// TIA Portal project "Network_1.0" (V15.1)

(* hardware
DEVICE "S71500/ET200MP station_1"  S7-1500 station
   slot 0: "Rail_0"  Rack  6ES7 590-1***0-0AA0
   slot 1: "PLC_1"  CPU 1516-3 PN/DP  6ES7 516-3AN01-0AB0  V2.6
      slot 3: "CPU display_1"  6ES7591-1BA00-0AA0
   slot 2: "AI 8xU/I/RTD/TC ST_1"  AI 8xU/I/RTD/TC ST  6ES7 531-7KF00-0AB0  V2.2
   slot 3: "AQ 4xU/I ST_1"  AQ 4xU/I ST  6ES7 532-5HD00-0AB0  V2.2
   slot 4: "DI 32x24VDC HF_1"  DI 32x24VDC HF  6ES7 521-1BL00-0AB0  V2.1
   slot 5: "DQ 32x24VDC/0.5A HF_1"  DQ 32x24VDC/0.5A HF  6ES7 522-1BL01-0AB0  V1.1
DEVICE "S7-1200 station_1"  S7-1200 Station
   slot 0: "Rack_0"  S7-1200 Rack  Rack  V1.0
   slot 1: "PLC_2"  CPU 1215C DC/DC/DC  6ES7 215-1AG40-0XB0  V4.2
DEVICE "S7-1200 station_2"  S7-1200 Station
   slot 0: "Rack_0"  S7-1200 Rack  Rack  V1.0
   slot 1: "PLC_3"  CPU 1215C DC/DC/DC  6ES7 215-1AG40-0XB0  V4.2
DEVICE "HMI_1"  KTP400 Basic PN
   slot 0: "HMI_1"  KTP400 Basic PN  6AV2 123-2DB03-0AX0  15.1.0.0
   slot 1: "HMI_RT_1"  KTP400 Basic PN  6AV2 123-2DB03-0AX0  15.1.0.0
   slot 5: "HMI_1.IE_CP_1"  PROFINET Interface  15.0.1.0
      slot 1: "PROFINET Interface_1"  PROFINET Interface
         slot 1: "Port_1"  Port
DEVICE "HMI_2"  KTP400 Basic PN
   slot 0: "HMI_2"  KTP400 Basic PN  6AV2 123-2DB03-0AX0  15.1.0.0
   slot 1: "HMI_RT_2"  KTP400 Basic PN  6AV2 123-2DB03-0AX0  15.1.0.0
   slot 5: "HMI_2.IE_CP_1"  PROFINET Interface  15.0.1.0
      slot 1: "PROFINET Interface_1"  PROFINET Interface
         slot 1: "Port_1"  Port
DEVICE "HMI_3"  KTP400 Basic PN
   slot 0: "HMI_3"  KTP400 Basic PN  6AV2 123-2DB03-0AX0  15.1.0.0
   slot 1: "HMI_RT_3"  KTP400 Basic PN  6AV2 123-2DB03-0AX0  15.1.0.0
   slot 5: "HMI_3.IE_CP_1"  PROFINET Interface  15.0.1.0
      slot 1: "PROFINET Interface_1"  PROFINET Interface
         slot 1: "Port_1"  Port
DEVICE "SCALANCE X005"  SCALANCE X-Station
   slot 0: "SCALANCE X rack"  Rail
   slot 0: "Switch_1"  6GK5 005-0BA00-1AB2  V1.0
*)

// ===== PLC "PLC_1"  CPU 1516-3 PN/DP =====

VAR_GLOBAL   // PLC tag table "Default tag table"
   "H2_Bet" AT %Q9.6 : Bool;
   "S1_Bet" AT %I17.4 : Bool;
   "S2_Bet" AT %I17.5 : Bool;
   "S3_Bet" AT %I17.6 : Bool;
   "S4_Bet" AT %I17.7 : Bool;
   "PE_Bet" AT %I17.3 : Bool;
   "H1_Bet" AT %Q9.5 : Bool;
   "H3_Bet" AT %Q9.7 : Bool;
   "Clock_Byte" AT %MB20 : Byte;
   "Clock_10Hz" AT %M20.0 : Bool;
   "Clock_5Hz" AT %M20.1 : Bool;
   "Clock_2.5Hz" AT %M20.2 : Bool;
   "Clock_2Hz" AT %M20.3 : Bool;
   "Clock_1.25Hz" AT %M20.4 : Bool;
   "Clock_1Hz" AT %M20.5 : Bool;
   "Clock_0.625Hz" AT %M20.6 : Bool;
   "Clock_0.5Hz" AT %M20.7 : Bool;
END_VAR

VAR_GLOBAL   // PLC tag table "PLC_1"
   "Selector_HMI_1" AT %MW8 : UInt;
   "Selector_HMI_2" AT %MW10 : UInt;
   "Selector_HMI_3" AT %MW12 : UInt;
   "S1_HM1" AT %M3.0 : Bool;
   "S2_HM1" AT %M3.1 : Bool;
   "S3_HM1" AT %M3.2 : Bool;
   "S1_HM2" AT %M3.3 : Bool;
   "S2_HM2" AT %M3.4 : Bool;
   "S3_HM2" AT %M3.5 : Bool;
   "S1_HM3" AT %M3.6 : Bool;
   "S2_HM3" AT %M3.7 : Bool;
   "S3_HM3" AT %M4.0 : Bool;
   "S1_PL1" AT %M4.1 : Bool;
   "S2_PL1" AT %M4.2 : Bool;
   "S3_PL1" AT %M4.3 : Bool;
   "S1_PL2" AT %M4.4 : Bool;
   "S2_PL2" AT %M4.5 : Bool;
   "S3_PL2" AT %M4.6 : Bool;
   "S1_PL3" AT %M4.7 : Bool;
   "S2_PL3" AT %M5.0 : Bool;
   "S3_PL3" AT %M5.1 : Bool;
   "H1_PL1" AT %M5.2 : Bool;
   "H2_PL1" AT %M5.3 : Bool;
   "H3_PL1" AT %M5.4 : Bool;
   "H1_PL2" AT %M5.5 : Bool;
   "H2_PL2" AT %M5.6 : Bool;
   "H3_PL2" AT %M5.7 : Bool;
   "H1_PL3" AT %M6.0 : Bool;
   "H2_PL3" AT %M6.1 : Bool;
   "H3_PL3" AT %M6.2 : Bool;
   "H1_HM1" AT %M6.3 : Bool;
   "H2_HM1" AT %M6.4 : Bool;
   "H3_HM1" AT %M6.5 : Bool;
   "H1_HM2" AT %M6.6 : Bool;
   "H2_HM2" AT %M6.7 : Bool;
   "H3_HM2" AT %M7.0 : Bool;
   "H1_HM3" AT %M7.1 : Bool;
   "H2_HM3" AT %M7.2 : Bool;
   "H3_HM3" AT %M7.3 : Bool;
END_VAR

DATA_BLOCK "COMS_PLC"   // DB1
{ S7_Optimized_Access := 'FALSE' }
VERSION : 0.1
   VAR
      PLC2_H1 : Int;
      PLC2_H2 : Int;
      PLC2_H3 : Int;
      PLC3_H1 : Int;
      PLC3_H2 : Int;
      PLC3_H3 : Int;
      PLC1_S1 : Int;
      PLC1_S2 : Int;
      PLC1_S3 : Int;
      PLC2_S1 : Int;
      PLC2_S2 : Int;
      PLC2_S3 : Int;
      PLC3_S1 : Int;
      PLC3_S2 : Int;
      PLC3_S3 : Int;
   END_VAR
BEGIN
END_DATA_BLOCK

ORGANIZATION_BLOCK "Main"   // OB1, LAD, ProgramCycle
TITLE = "Main Program Sweep (Cycle)"
{ S7_Optimized_Access := 'TRUE' }
VERSION : 0.1
   VAR_INPUT
      Initial_Call : Bool;   // Initial call of this OB
      Remanence : Bool;   // =True, if remanent data are available
   END_VAR
BEGIN

REGION Network 1: Salidas a HMI1
   // Salidas a HMI Selector 1
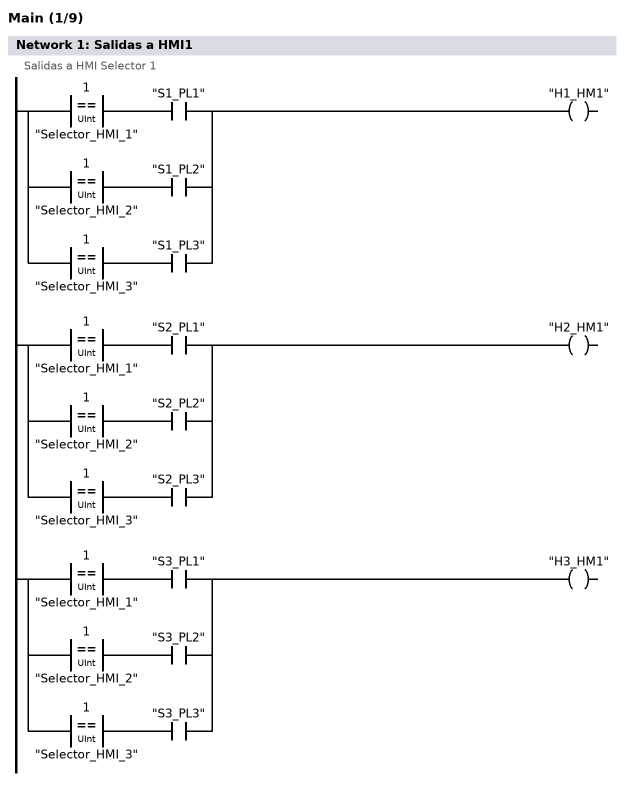
   RUNG wire#powerrail
      { S7_Templates := "SrcType := UInt" } EQ_Contact(in1 := 1, in2 := "Selector_HMI_1")
      Contact( "S1_PL1" )
      wire#w1
      Coil( "H1_HM1" )
   END_RUNG
   RUNG wire#powerrail
      { S7_Templates := "SrcType := UInt" } EQ_Contact(in1 := 1, in2 := "Selector_HMI_2")
      Contact( "S1_PL2" )
   END_RUNG wire#w1
   RUNG wire#powerrail
      { S7_Templates := "SrcType := UInt" } EQ_Contact(in1 := 1, in2 := "Selector_HMI_3")
      Contact( "S1_PL3" )
   END_RUNG wire#w1
   RUNG wire#powerrail
      { S7_Templates := "SrcType := UInt" } EQ_Contact(in1 := 1, in2 := "Selector_HMI_1")
      Contact( "S2_PL1" )
      wire#w2
      Coil( "H2_HM1" )
   END_RUNG
   RUNG wire#powerrail
      { S7_Templates := "SrcType := UInt" } EQ_Contact(in1 := 1, in2 := "Selector_HMI_2")
      Contact( "S2_PL2" )
   END_RUNG wire#w2
   RUNG wire#powerrail
      { S7_Templates := "SrcType := UInt" } EQ_Contact(in1 := 1, in2 := "Selector_HMI_3")
      Contact( "S2_PL3" )
   END_RUNG wire#w2
   RUNG wire#powerrail
      { S7_Templates := "SrcType := UInt" } EQ_Contact(in1 := 1, in2 := "Selector_HMI_1")
      Contact( "S3_PL1" )
      wire#w3
      Coil( "H3_HM1" )
   END_RUNG
   RUNG wire#powerrail
      { S7_Templates := "SrcType := UInt" } EQ_Contact(in1 := 1, in2 := "Selector_HMI_2")
      Contact( "S3_PL2" )
   END_RUNG wire#w3
   RUNG wire#powerrail
      { S7_Templates := "SrcType := UInt" } EQ_Contact(in1 := 1, in2 := "Selector_HMI_3")
      Contact( "S3_PL3" )
   END_RUNG wire#w3
   // the same network as SCL:
   "H1_HM1" := ((1 = "Selector_HMI_1") AND "S1_PL1") OR ((1 = "Selector_HMI_2") AND "S1_PL2") OR ((1 = "Selector_HMI_3") AND "S1_PL3");
   "H2_HM1" := ((1 = "Selector_HMI_1") AND "S2_PL1") OR ((1 = "Selector_HMI_2") AND "S2_PL2") OR ((1 = "Selector_HMI_3") AND "S2_PL3");
   "H3_HM1" := ((1 = "Selector_HMI_1") AND "S3_PL1") OR ((1 = "Selector_HMI_2") AND "S3_PL2") OR ((1 = "Selector_HMI_3") AND "S3_PL3");
END_REGION

REGION Network 2: Salidas a HMI2
   // Salidas a HMI Selector 1
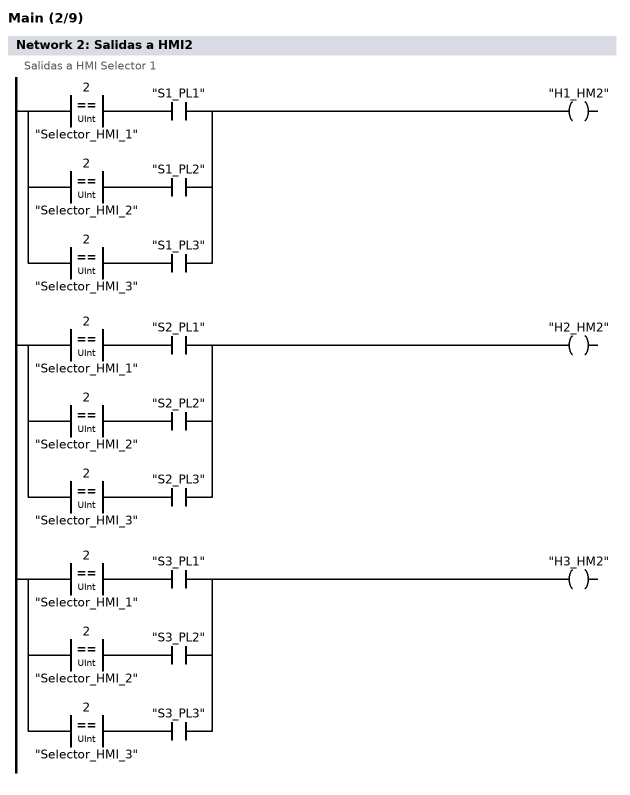
   RUNG wire#powerrail
      { S7_Templates := "SrcType := UInt" } EQ_Contact(in1 := 2, in2 := "Selector_HMI_1")
      Contact( "S1_PL1" )
      wire#w1
      Coil( "H1_HM2" )
   END_RUNG
   RUNG wire#powerrail
      { S7_Templates := "SrcType := UInt" } EQ_Contact(in1 := 2, in2 := "Selector_HMI_2")
      Contact( "S1_PL2" )
   END_RUNG wire#w1
   RUNG wire#powerrail
      { S7_Templates := "SrcType := UInt" } EQ_Contact(in1 := 2, in2 := "Selector_HMI_3")
      Contact( "S1_PL3" )
   END_RUNG wire#w1
   RUNG wire#powerrail
      { S7_Templates := "SrcType := UInt" } EQ_Contact(in1 := 2, in2 := "Selector_HMI_1")
      Contact( "S2_PL1" )
      wire#w2
      Coil( "H2_HM2" )
   END_RUNG
   RUNG wire#powerrail
      { S7_Templates := "SrcType := UInt" } EQ_Contact(in1 := 2, in2 := "Selector_HMI_2")
      Contact( "S2_PL2" )
   END_RUNG wire#w2
   RUNG wire#powerrail
      { S7_Templates := "SrcType := UInt" } EQ_Contact(in1 := 2, in2 := "Selector_HMI_3")
      Contact( "S2_PL3" )
   END_RUNG wire#w2
   RUNG wire#powerrail
      { S7_Templates := "SrcType := UInt" } EQ_Contact(in1 := 2, in2 := "Selector_HMI_1")
      Contact( "S3_PL1" )
      wire#w3
      Coil( "H3_HM2" )
   END_RUNG
   RUNG wire#powerrail
      { S7_Templates := "SrcType := UInt" } EQ_Contact(in1 := 2, in2 := "Selector_HMI_2")
      Contact( "S3_PL2" )
   END_RUNG wire#w3
   RUNG wire#powerrail
      { S7_Templates := "SrcType := UInt" } EQ_Contact(in1 := 2, in2 := "Selector_HMI_3")
      Contact( "S3_PL3" )
   END_RUNG wire#w3
   // the same network as SCL:
   "H1_HM2" := ((2 = "Selector_HMI_1") AND "S1_PL1") OR ((2 = "Selector_HMI_2") AND "S1_PL2") OR ((2 = "Selector_HMI_3") AND "S1_PL3");
   "H2_HM2" := ((2 = "Selector_HMI_1") AND "S2_PL1") OR ((2 = "Selector_HMI_2") AND "S2_PL2") OR ((2 = "Selector_HMI_3") AND "S2_PL3");
   "H3_HM2" := ((2 = "Selector_HMI_1") AND "S3_PL1") OR ((2 = "Selector_HMI_2") AND "S3_PL2") OR ((2 = "Selector_HMI_3") AND "S3_PL3");
END_REGION

REGION Network 3: Salidas a HMI3
   // Salidas a HMI Selector 1
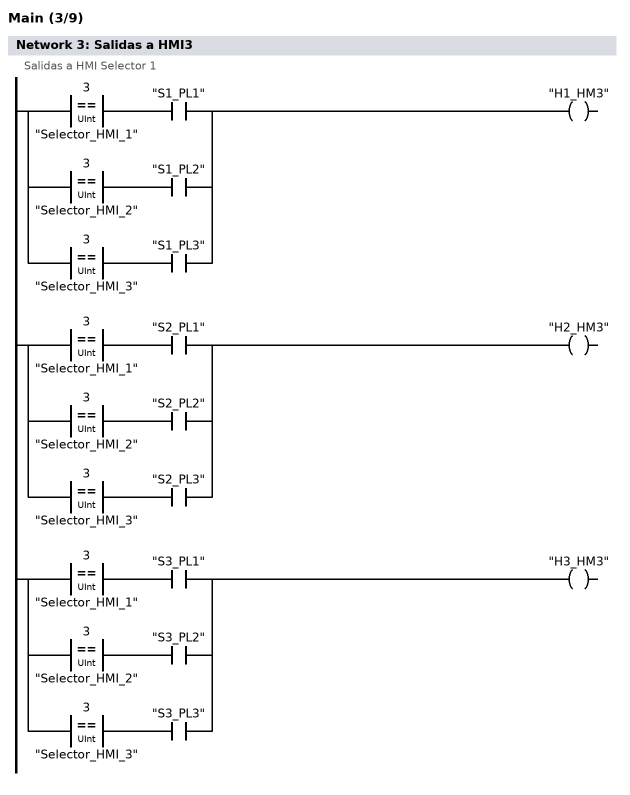
   RUNG wire#powerrail
      { S7_Templates := "SrcType := UInt" } EQ_Contact(in1 := 3, in2 := "Selector_HMI_1")
      Contact( "S1_PL1" )
      wire#w1
      Coil( "H1_HM3" )
   END_RUNG
   RUNG wire#powerrail
      { S7_Templates := "SrcType := UInt" } EQ_Contact(in1 := 3, in2 := "Selector_HMI_2")
      Contact( "S1_PL2" )
   END_RUNG wire#w1
   RUNG wire#powerrail
      { S7_Templates := "SrcType := UInt" } EQ_Contact(in1 := 3, in2 := "Selector_HMI_3")
      Contact( "S1_PL3" )
   END_RUNG wire#w1
   RUNG wire#powerrail
      { S7_Templates := "SrcType := UInt" } EQ_Contact(in1 := 3, in2 := "Selector_HMI_1")
      Contact( "S2_PL1" )
      wire#w2
      Coil( "H2_HM3" )
   END_RUNG
   RUNG wire#powerrail
      { S7_Templates := "SrcType := UInt" } EQ_Contact(in1 := 3, in2 := "Selector_HMI_2")
      Contact( "S2_PL2" )
   END_RUNG wire#w2
   RUNG wire#powerrail
      { S7_Templates := "SrcType := UInt" } EQ_Contact(in1 := 3, in2 := "Selector_HMI_3")
      Contact( "S2_PL3" )
   END_RUNG wire#w2
   RUNG wire#powerrail
      { S7_Templates := "SrcType := UInt" } EQ_Contact(in1 := 3, in2 := "Selector_HMI_1")
      Contact( "S3_PL1" )
      wire#w3
      Coil( "H3_HM3" )
   END_RUNG
   RUNG wire#powerrail
      { S7_Templates := "SrcType := UInt" } EQ_Contact(in1 := 3, in2 := "Selector_HMI_2")
      Contact( "S3_PL2" )
   END_RUNG wire#w3
   RUNG wire#powerrail
      { S7_Templates := "SrcType := UInt" } EQ_Contact(in1 := 3, in2 := "Selector_HMI_3")
      Contact( "S3_PL3" )
   END_RUNG wire#w3
   // the same network as SCL:
   "H1_HM3" := ((3 = "Selector_HMI_1") AND "S1_PL1") OR ((3 = "Selector_HMI_2") AND "S1_PL2") OR ((3 = "Selector_HMI_3") AND "S1_PL3");
   "H2_HM3" := ((3 = "Selector_HMI_1") AND "S2_PL1") OR ((3 = "Selector_HMI_2") AND "S2_PL2") OR ((3 = "Selector_HMI_3") AND "S2_PL3");
   "H3_HM3" := ((3 = "Selector_HMI_1") AND "S3_PL1") OR ((3 = "Selector_HMI_2") AND "S3_PL2") OR ((3 = "Selector_HMI_3") AND "S3_PL3");
END_REGION

REGION Network 4: Salidas a PLC1
   // Salidas a HMI Selector 1
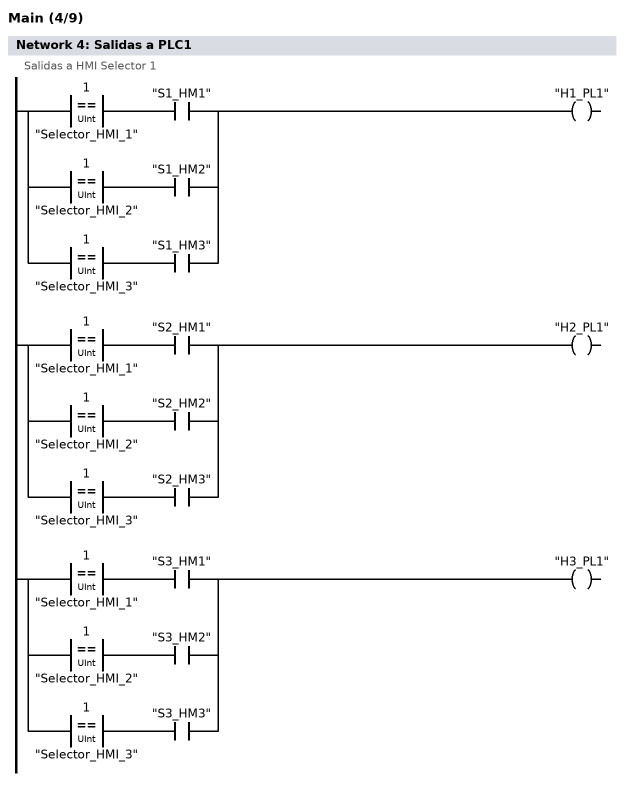
   RUNG wire#powerrail
      { S7_Templates := "SrcType := UInt" } EQ_Contact(in1 := 1, in2 := "Selector_HMI_1")
      Contact( "S1_HM1" )
      wire#w1
      Coil( "H1_PL1" )
   END_RUNG
   RUNG wire#powerrail
      { S7_Templates := "SrcType := UInt" } EQ_Contact(in1 := 1, in2 := "Selector_HMI_2")
      Contact( "S1_HM2" )
   END_RUNG wire#w1
   RUNG wire#powerrail
      { S7_Templates := "SrcType := UInt" } EQ_Contact(in1 := 1, in2 := "Selector_HMI_3")
      Contact( "S1_HM3" )
   END_RUNG wire#w1
   RUNG wire#powerrail
      { S7_Templates := "SrcType := UInt" } EQ_Contact(in1 := 1, in2 := "Selector_HMI_1")
      Contact( "S2_HM1" )
      wire#w2
      Coil( "H2_PL1" )
   END_RUNG
   RUNG wire#powerrail
      { S7_Templates := "SrcType := UInt" } EQ_Contact(in1 := 1, in2 := "Selector_HMI_2")
      Contact( "S2_HM2" )
   END_RUNG wire#w2
   RUNG wire#powerrail
      { S7_Templates := "SrcType := UInt" } EQ_Contact(in1 := 1, in2 := "Selector_HMI_3")
      Contact( "S2_HM3" )
   END_RUNG wire#w2
   RUNG wire#powerrail
      { S7_Templates := "SrcType := UInt" } EQ_Contact(in1 := 1, in2 := "Selector_HMI_1")
      Contact( "S3_HM1" )
      wire#w3
      Coil( "H3_PL1" )
   END_RUNG
   RUNG wire#powerrail
      { S7_Templates := "SrcType := UInt" } EQ_Contact(in1 := 1, in2 := "Selector_HMI_2")
      Contact( "S3_HM2" )
   END_RUNG wire#w3
   RUNG wire#powerrail
      { S7_Templates := "SrcType := UInt" } EQ_Contact(in1 := 1, in2 := "Selector_HMI_3")
      Contact( "S3_HM3" )
   END_RUNG wire#w3
   // the same network as SCL:
   "H1_PL1" := ((1 = "Selector_HMI_1") AND "S1_HM1") OR ((1 = "Selector_HMI_2") AND "S1_HM2") OR ((1 = "Selector_HMI_3") AND "S1_HM3");
   "H2_PL1" := ((1 = "Selector_HMI_1") AND "S2_HM1") OR ((1 = "Selector_HMI_2") AND "S2_HM2") OR ((1 = "Selector_HMI_3") AND "S2_HM3");
   "H3_PL1" := ((1 = "Selector_HMI_1") AND "S3_HM1") OR ((1 = "Selector_HMI_2") AND "S3_HM2") OR ((1 = "Selector_HMI_3") AND "S3_HM3");
END_REGION

REGION Network 5: Salidas a PLC2
   // Salidas a HMI Selector 1
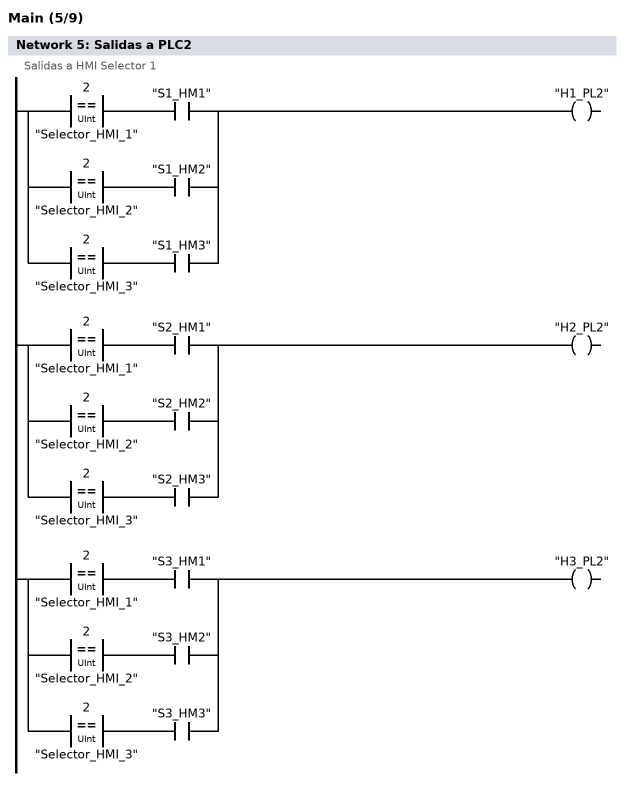
   RUNG wire#powerrail
      { S7_Templates := "SrcType := UInt" } EQ_Contact(in1 := 2, in2 := "Selector_HMI_1")
      Contact( "S1_HM1" )
      wire#w1
      Coil( "H1_PL2" )
   END_RUNG
   RUNG wire#powerrail
      { S7_Templates := "SrcType := UInt" } EQ_Contact(in1 := 2, in2 := "Selector_HMI_2")
      Contact( "S1_HM2" )
   END_RUNG wire#w1
   RUNG wire#powerrail
      { S7_Templates := "SrcType := UInt" } EQ_Contact(in1 := 2, in2 := "Selector_HMI_3")
      Contact( "S1_HM3" )
   END_RUNG wire#w1
   RUNG wire#powerrail
      { S7_Templates := "SrcType := UInt" } EQ_Contact(in1 := 2, in2 := "Selector_HMI_1")
      Contact( "S2_HM1" )
      wire#w2
      Coil( "H2_PL2" )
   END_RUNG
   RUNG wire#powerrail
      { S7_Templates := "SrcType := UInt" } EQ_Contact(in1 := 2, in2 := "Selector_HMI_2")
      Contact( "S2_HM2" )
   END_RUNG wire#w2
   RUNG wire#powerrail
      { S7_Templates := "SrcType := UInt" } EQ_Contact(in1 := 2, in2 := "Selector_HMI_3")
      Contact( "S2_HM3" )
   END_RUNG wire#w2
   RUNG wire#powerrail
      { S7_Templates := "SrcType := UInt" } EQ_Contact(in1 := 2, in2 := "Selector_HMI_1")
      Contact( "S3_HM1" )
      wire#w3
      Coil( "H3_PL2" )
   END_RUNG
   RUNG wire#powerrail
      { S7_Templates := "SrcType := UInt" } EQ_Contact(in1 := 2, in2 := "Selector_HMI_2")
      Contact( "S3_HM2" )
   END_RUNG wire#w3
   RUNG wire#powerrail
      { S7_Templates := "SrcType := UInt" } EQ_Contact(in1 := 2, in2 := "Selector_HMI_3")
      Contact( "S3_HM3" )
   END_RUNG wire#w3
   // the same network as SCL:
   "H1_PL2" := ((2 = "Selector_HMI_1") AND "S1_HM1") OR ((2 = "Selector_HMI_2") AND "S1_HM2") OR ((2 = "Selector_HMI_3") AND "S1_HM3");
   "H2_PL2" := ((2 = "Selector_HMI_1") AND "S2_HM1") OR ((2 = "Selector_HMI_2") AND "S2_HM2") OR ((2 = "Selector_HMI_3") AND "S2_HM3");
   "H3_PL2" := ((2 = "Selector_HMI_1") AND "S3_HM1") OR ((2 = "Selector_HMI_2") AND "S3_HM2") OR ((2 = "Selector_HMI_3") AND "S3_HM3");
END_REGION

REGION Network 6: Salidas a PLC3
   // Salidas a HMI Selector 1
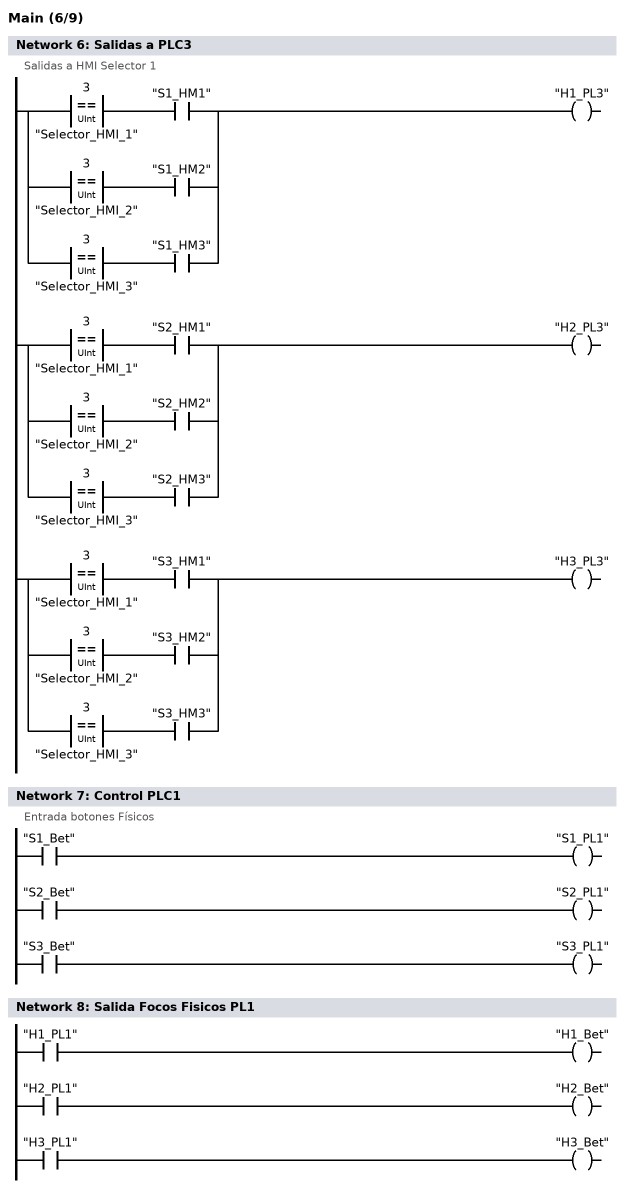
   RUNG wire#powerrail
      { S7_Templates := "SrcType := UInt" } EQ_Contact(in1 := 3, in2 := "Selector_HMI_1")
      Contact( "S1_HM1" )
      wire#w1
      Coil( "H1_PL3" )
   END_RUNG
   RUNG wire#powerrail
      { S7_Templates := "SrcType := UInt" } EQ_Contact(in1 := 3, in2 := "Selector_HMI_2")
      Contact( "S1_HM2" )
   END_RUNG wire#w1
   RUNG wire#powerrail
      { S7_Templates := "SrcType := UInt" } EQ_Contact(in1 := 3, in2 := "Selector_HMI_3")
      Contact( "S1_HM3" )
   END_RUNG wire#w1
   RUNG wire#powerrail
      { S7_Templates := "SrcType := UInt" } EQ_Contact(in1 := 3, in2 := "Selector_HMI_1")
      Contact( "S2_HM1" )
      wire#w2
      Coil( "H2_PL3" )
   END_RUNG
   RUNG wire#powerrail
      { S7_Templates := "SrcType := UInt" } EQ_Contact(in1 := 3, in2 := "Selector_HMI_2")
      Contact( "S2_HM2" )
   END_RUNG wire#w2
   RUNG wire#powerrail
      { S7_Templates := "SrcType := UInt" } EQ_Contact(in1 := 3, in2 := "Selector_HMI_3")
      Contact( "S2_HM3" )
   END_RUNG wire#w2
   RUNG wire#powerrail
      { S7_Templates := "SrcType := UInt" } EQ_Contact(in1 := 3, in2 := "Selector_HMI_1")
      Contact( "S3_HM1" )
      wire#w3
      Coil( "H3_PL3" )
   END_RUNG
   RUNG wire#powerrail
      { S7_Templates := "SrcType := UInt" } EQ_Contact(in1 := 3, in2 := "Selector_HMI_2")
      Contact( "S3_HM2" )
   END_RUNG wire#w3
   RUNG wire#powerrail
      { S7_Templates := "SrcType := UInt" } EQ_Contact(in1 := 3, in2 := "Selector_HMI_3")
      Contact( "S3_HM3" )
   END_RUNG wire#w3
   // the same network as SCL:
   "H1_PL3" := ((3 = "Selector_HMI_1") AND "S1_HM1") OR ((3 = "Selector_HMI_2") AND "S1_HM2") OR ((3 = "Selector_HMI_3") AND "S1_HM3");
   "H2_PL3" := ((3 = "Selector_HMI_1") AND "S2_HM1") OR ((3 = "Selector_HMI_2") AND "S2_HM2") OR ((3 = "Selector_HMI_3") AND "S2_HM3");
   "H3_PL3" := ((3 = "Selector_HMI_1") AND "S3_HM1") OR ((3 = "Selector_HMI_2") AND "S3_HM2") OR ((3 = "Selector_HMI_3") AND "S3_HM3");
END_REGION

REGION Network 7: Control PLC1
   // Entrada botones Físicos
   RUNG wire#powerrail
      Contact( "S1_Bet" )
      Coil( "S1_PL1" )
   END_RUNG
   RUNG wire#powerrail
      Contact( "S2_Bet" )
      Coil( "S2_PL1" )
   END_RUNG
   RUNG wire#powerrail
      Contact( "S3_Bet" )
      Coil( "S3_PL1" )
   END_RUNG
   // the same network as SCL:
   "S1_PL1" := "S1_Bet";
   "S2_PL1" := "S2_Bet";
   "S3_PL1" := "S3_Bet";
END_REGION

REGION Network 8: Salida Focos Fisicos PL1
   RUNG wire#powerrail
      Contact( "H1_PL1" )
      Coil( "H1_Bet" )
   END_RUNG
   RUNG wire#powerrail
      Contact( "H2_PL1" )
      Coil( "H2_Bet" )
   END_RUNG
   RUNG wire#powerrail
      Contact( "H3_PL1" )
      Coil( "H3_Bet" )
   END_RUNG
   // the same network as SCL:
   "H1_Bet" := "H1_PL1";
   "H2_Bet" := "H2_PL1";
   "H3_Bet" := "H3_PL1";
END_REGION

REGION Network 9: LECTURAS PLC
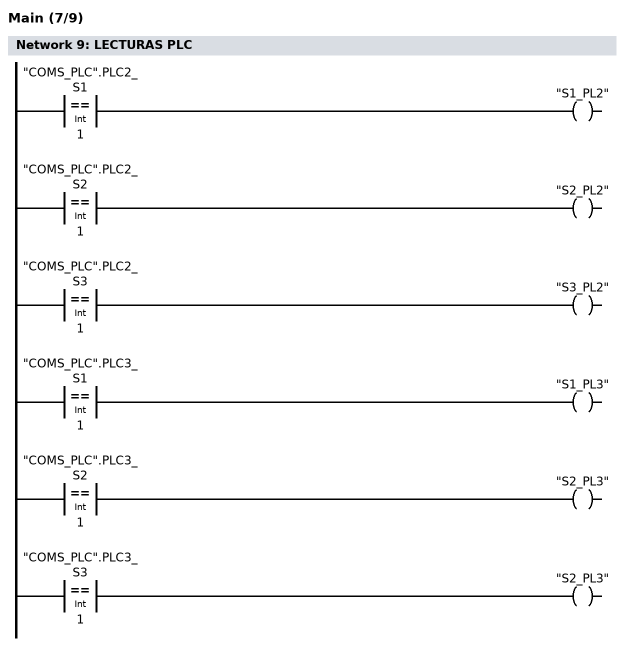
   RUNG wire#powerrail
      { S7_Templates := "SrcType := Int" } EQ_Contact(in1 := "COMS_PLC".PLC2_S1, in2 := 1)
      Coil( "S1_PL2" )
   END_RUNG
   RUNG wire#powerrail
      { S7_Templates := "SrcType := Int" } EQ_Contact(in1 := "COMS_PLC".PLC2_S2, in2 := 1)
      Coil( "S2_PL2" )
   END_RUNG
   RUNG wire#powerrail
      { S7_Templates := "SrcType := Int" } EQ_Contact(in1 := "COMS_PLC".PLC2_S3, in2 := 1)
      Coil( "S3_PL2" )
   END_RUNG
   RUNG wire#powerrail
      { S7_Templates := "SrcType := Int" } EQ_Contact(in1 := "COMS_PLC".PLC3_S1, in2 := 1)
      Coil( "S1_PL3" )
   END_RUNG
   RUNG wire#powerrail
      { S7_Templates := "SrcType := Int" } EQ_Contact(in1 := "COMS_PLC".PLC3_S2, in2 := 1)
      Coil( "S2_PL3" )
   END_RUNG
   RUNG wire#powerrail
      { S7_Templates := "SrcType := Int" } EQ_Contact(in1 := "COMS_PLC".PLC3_S3, in2 := 1)
      Coil( "S2_PL3" )
   END_RUNG
   // the same network as SCL:
   "S1_PL2" := "COMS_PLC".PLC2_S1 = 1;
   "S2_PL2" := "COMS_PLC".PLC2_S2 = 1;
   "S3_PL2" := "COMS_PLC".PLC2_S3 = 1;
   "S1_PL3" := "COMS_PLC".PLC3_S1 = 1;
   "S2_PL3" := "COMS_PLC".PLC3_S2 = 1;
   "S2_PL3" := "COMS_PLC".PLC3_S3 = 1;
END_REGION

REGION Network 10: INSERT DB